VERSION : 0.1
   STRUCT
      dMissionCode : DInt;   // Mission code number
      rgdFireHeadThreshold_cmm : Array[0.."CONST_dNumberOfHeadsCycle"] of DInt;   // Head#x firing threshold [mm/100]
      rgdHeadsPositions_cmm : Array[0.."CONST_dNumberOfHeadsCycle"] of DInt;   // Head#x positions request [mm/100]
      rgxFireHeadON_OFF : Array[0.."CONST_dNumberOfHeadsCycle"] of Bool;   // Head#x firing type request [bit]
      rgxDataToProcessInter : Array[0.."CONST_dNumberOfHeadsCycle"] of Bool;   // Head#x data to process by interrupt
      xGateOpen : Bool;   // Interrupt gate open
      dTargetLineValue_cmm : DInt;   // Virtual target line value [mm/100]
      rgxArmRequest : Array[0.."CONST_dNumberOfHeadsCycle"] of Bool;   // Head#x arming request
      rgdArmRequestTarget_cmm : Array[0.."CONST_dNumberOfHeadsCycle"] of DInt;   // Arm request target virtual [mm/100]
      rgxOilRequest : Array[0.."CONST_dNumberOfHeadsCycle"] of Bool;   // Head#x oil request
      rgdOilRequestTarget_cmm : Array[0.."CONST_dNumberOfHeadsCycle"] of DInt;   // Oil request target virtual [mm/100]
      rgdArmRequestIDMission : Array[0.."CONST_dNumberOfHeadsCycle"] of DInt;   // Arm request ID mission
      rgdOilRequestIDMission : Array[0.."CONST_dNumberOfHeadsCycle"] of DInt;   // Oil request ID mission
   END_STRUCT;
END_TYPE

TYPE "UDT_DataManager_Tank"
VERSION : 0.1
   STRUCT
      dMissionCode : DInt;   // Mission code
      dMissionValue_cmm : DInt;   // Mission value [mm/100]
      rgxFireRequest : Array[0.."CONST_dNumberOfHeadsCycle"] of Bool;   // Head#x fire request
      rgdHeadsPositions_cmm : Array[0.."CONST_dNumberOfHeadsCycle"] of DInt;   // Head#x position request [mm/100]
   END_STRUCT;
END_TYPE

TYPE "UDT_MB_ConnData"
   STRUCT
      IP_OCTET_1 : USInt;
      IP_OCTET_2 : USInt;
      IP_OCTET_3 : USInt;
      IP_OCTET_4 : USInt;
      ConnectID1 : Conn_Ouc;
      ConnectID2 : Conn_Ouc;
      ConnectID3 : Conn_Ouc;
      ConnectID4 : Conn_Ouc;
   END_STRUCT;
END_TYPE

TYPE "UDT_CM_IDEV_FromMainLine"
VERSION : 0.1
   STRUCT
      dSpare1 : Array[0..2] of DInt;
      xCycleON : Bool;   // Cycle ON
      xResetAnomaly : Bool;   // Reset anomaly
      xResetBuffers : Bool;   // Reset buffer
      xGlassBreak : Bool;   // Glass break under the bridge
      xPLCActive0 : Bool;   // PLC Active (0=CPU0, 1=CPU1)
      xPLCActive1 : Bool;   // PLC Active (0=CPU0, 1=CPU1)
      xQLTplate : Bool;   // Quality plate in progress
      xSpare2 : Bool;
      xSpare3 : Bool;
      xSpare4 : Bool;
      xSpare5 : Bool;
      xSpare6 : Bool;
      xSpare7 : Bool;
      xSpare8 : Bool;
      xSpare9 : Bool;
      xSpare10 : Bool;
      xStatusSpare : Array[0..15] of Bool;
      dSpare2 : Array[0..7] of DInt;
      iSpare : Int;
   END_STRUCT;
END_TYPE

TYPE "UDT_CM_IDEV_ToMainLine"
VERSION : 0.1
   STRUCT
      dProcessingIDPlate : DInt;   // Processing ID Plate [Num]
      dSpare1 : DInt;
      dSpare2 : DInt;
      rgxStatus : Array[0..31] of Bool;   // Status heads
      rgdHeadsPositions_cmm : Array[0..15] of DInt;   // Head #x position status
      rgxHeadStatus : Array[0..15] of Bool;   // Head #x enabled
      rgxCuttingStatus : Array[0..15] of Bool;   // Head #x cuuting status
      rgdHeadsPressure : Array[0..15] of DInt;   // Head #x Pressure [mN]
      rgrHeadsSpace : Array[0..15] of Real;   // Head #x Distance [Km]
      iFireOffset_ON : Int;   // All head fire on offset
      iFireOffset_OFF : Int;   // All head fire off offset
      iSpare : Int;
      dSpare : Array[0..7] of DInt;
   END_STRUCT;
   // // rgxStatus[0] : Glass break in progress
   // // rgxStatus[1] : Liftup pushbutton engaged
   // // rgxStatus[2] : Bridge enabled
   // // rgxStatus[3] : Bridge locked
   // // rgxStatus[8] : Fire offset calibration
END_TYPE

TYPE "UDT_CM_RECV_SyncroData"
VERSION : 0.1
   STRUCT
      dMissionID : DInt;   // Mission Identifier
      dSynchroValue_cmm : DInt;   // Counter value in the last synchro [mm/100]
      dSpare : Array[0..7] of DInt;
      xSpare : Array[0..15] of Bool;
      dSpare2 : Array[0..2] of DInt;
      iSpare : Int;
   END_STRUCT;
END_TYPE

TYPE "UDT_CM_RECV_MissionData"
VERSION : 0.1
   STRUCT
      dMissionID : DInt;   // Mission Identifier
      dMissionStart_cmm : DInt;   // Mission counter start [mm/100]
      dMissionEnd_cmm : DInt;   // Mission counter stop [mm/100]
      dTrackingDbNumber : DInt;   // Tracking DB number
      dSpare1 : Array[0..9] of DInt;
      rgxFireRequest : Array[0..31] of Bool;   // Head #x firing request
      rgdHeadsPosition_cmm : Array[0..15] of DInt;   // Head #x position request [mm/100]
      dSpare2 : Array[0..14] of DInt;
   END_STRUCT;
END_TYPE

TYPE "UDT_CM_Manager"
VERSION : 0.1
   STRUCT
      ST_xNewDataReceiveCPU0 : Bool;   // New data receive
      ST_xErrorCPU0 : Bool;   // Error
      ST_xNewSynchCPU0 : Bool;   // New synch
      ST_xNewMissionCPU0 : Bool;   // New mission
      AUX_iDataLenghtCPU0 : Word;   // Data lenght
      AUX_iStateCPU0 : Int;   // Status
      ST_xNewDataReceiveCPU1 : Bool;   // New data receive
      ST_xErrorCPU1 : Bool;   // Error
      ST_xNewSynchCPU1 : Bool;   // New synch
      ST_xNewMissionCPU1 : Bool;   // New mission
      AUX_iDataLenghtCPU1 : Word;   // Data lenght
      AUX_iStateCPU1 : Int;   // Status
      AUX_tmON_ConsumedTimeout : IEC_TIMER;   // Timer ON consumed timeout PLCA
      AUX_rgdHeadMissionIDInProg_Copy : Array[0.."CONST_dNumberOfHeadsCycle"] of DInt;   // Head#x mission ID in progress
      AUX_rgxHeadFiringMissionInProg_Copy : Array[0.."CONST_dNumberOfHeadsCycle"] of Bool;   // Head#x firing mission in progress
      ST_xConsumedTimeout : Bool;   // Consumed message timeout PLCA
      ST_xMissionPacketLost : Bool;   // Mission message packet lost PLC A
      ST_xSyncroPacketLost : Bool;   // Syncro message packet lost PLC A
      ST_MutingFiringOB : Bool;   // Muting Ob30 firing
   END_STRUCT;
END_TYPE

TYPE "UDT_HeadPar"
VERSION : 0.1
   STRUCT
      iAddress : Int;
      iLength : Byte;
      dValue : DInt;
   END_STRUCT;
END_TYPE

TYPE "UDT_AxisParameters"
VERSION : 0.1
   STRUCT
      rgtAxisParameters : Array[0..20] of "UDT_HeadPar";
      dParametersToDownload : DInt;
   END_STRUCT;
END_TYPE

TYPE "UDT_BRCV_FromMainLine"
VERSION : 0.1
   STRUCT
      SyncroData : "UDT_CM_RECV_SyncroData";
      MissionData : "UDT_CM_RECV_MissionData";
   END_STRUCT;
END_TYPE

TYPE "LPD_typeCountFeedbackCh"
VERSION : 0.1
   STRUCT
      countValue : DInt := 16#0000;   // Current count value
      capturedValue : DInt := 16#0000;   // Last Capture value acquired
      measuredValue : Real := 0.0;   // Current measured value
      powerError : Bool := FALSE;   // Incorrect supply voltage L+
      encError : Bool := FALSE;   // Incorrect encoder signal
      ldError : Bool := FALSE;   // Error when loading via control interface
      reserved1 : Bool := FALSE;   // Reserved
      reserved2 : Bool := FALSE;   // Reserved
      reserved3 : Bool := FALSE;   // Reserved
      reserved4 : Bool := FALSE;   // Reserved
      reserved5 : Bool := FALSE;   // Reserved
      commActive : Bool := FALSE;   // Comm active
      resEventAck : Bool := FALSE;   // Reset of event bits active
      ldStsSlot0 : Bool := FALSE;   // Load request for Slot 0 detected and executed (toggling)
      ldStsSlot1 : Bool := FALSE;   // Load request for Slot 1 detected and executed (toggling)
      stsReady : Bool := FALSE;   // Digital on-board I/O started up and parameters assigned
      stsSwGate : Bool := FALSE;   // Software gate status
      reserved7 : Bool := FALSE;   // Reserved
      reserved8 : Bool := FALSE;   // Reserved
      stsDir : Bool := FALSE;   // Direction of last count value change
      stsCount : Bool := FALSE;   // Count pulse detected within last approx. 0.5 s
      stsGate : Bool := FALSE;   // Internal gate status
      stsDQ0 : Bool := FALSE;   // Status HSC DQ0
      stsDQ1 : Bool := FALSE;   // Status HSC DQ1
      stsDI0 : Bool := FALSE;   // Status HSC DI0
      stsDI1 : Bool := FALSE;   // Status HSC DI1
      stsDI2 : Bool := FALSE;   // Status HSC DI2
      eventZero : Bool := FALSE;   // Zero crossing has occurred
      eventUnderflow : Bool := FALSE;   // Underflow has occurred
      eventOverflow : Bool := FALSE;   // Overflow has occurred
      eventCompare0 : Bool := FALSE;   // Comparison event for DQ0 has occurred
      eventCompare1 : Bool := FALSE;   // Comparison event for DQ1 has occurred
      eventSync : Bool := FALSE;   // Synchronization has occurred
      eventCapture : Bool := FALSE;   // Capture event has occurred
      stsMeasInterval : Bool := FALSE;   // Count pulse detected in previous measuring interval
   END_STRUCT;
END_TYPE

TYPE "LPD_typeCountControlCh"
VERSION : 0.1
   STRUCT
      loadValue0 : DWord := 16#0000;   // Load value 0
      loadValue1 : DWord := 16#0000;   // Load value 1
      controlByte : Byte := B#16#00;   // Control byte load value
      swGate : Bool := FALSE;   // Software gate
      tmCtrlDQ0 : Bool := FALSE;   // Enable technological function DQ0
      tmCtrlDQ1 : Bool := FALSE;   // Enable technological function DQ1
      setDQ0 : Bool := FALSE;   // Set DQ0
      setDQ1 : Bool := FALSE;   // Set DQ1
      enSyncUp : Bool := FALSE;   // Enable upward synchronization
      enSyncDown : Bool := FALSE;   // Enable downward synchronization
      enCapture : Bool := FALSE;   // Enable capture function
      resError : Bool := FALSE;   // Reset of saved error states
      resEvent : Bool := FALSE;   // Reset of saved events
      reserved0 : Bool := FALSE;   // Reserved
      reserved1 : Bool := FALSE;   // Reserved
      reserved2 : Bool := FALSE;   // Reserved
      reserved3 : Bool := FALSE;   // Reserved
      reserved4 : Bool := FALSE;   // Reserved
      SetDir : Bool := FALSE;   // Count direction (with encoder without direction signal)
      reserved5 : Byte;   // Reserved
   END_STRUCT;
END_TYPE

// folder: ProfinetDiagnostic

TYPE "TINFO_"
VERSION : 0.1
   STRUCT
      OB_start_info : Array[0..19] of Byte;
      W_20_STATION : Word;
      B22_slave_type : Byte;
      B23_interrupt_type : Byte;
      B24_origination : Byte;
      B25_diag_flag : Byte;
      W26_PN_ID : Word;
      W28_MFG_ID : Word;
      W30_INST_ID : Word;
      other_data : Array[1..70] of Byte;
   END_STRUCT;
END_TYPE

TYPE "AINFO_"
VERSION : 0.1
   STRUCT
      W0_block_type : Word;
      W2_block_length : Word;
      W4_version : Word;
      W6_interrupt_type : Word;
      D8_API : DWord;
      W12_comp_slot_num : Word;
      W14_submodule_slot_num : Word;
      D16_module_ID : DWord;
      D20_submodule_ID : DWord;
      W24_interrupt_specifer : Word;
      Add_W0_format_ID : Word;
      Add_W2_channel_num : Word;
      Add_B4_error_info : Byte;
      Add_B5_data_format : Byte;
      Add_W6_error_type : Word;
      extended_info : Array[34..1431] of Byte;
   END_STRUCT;
END_TYPE

TYPE "PN_Alarm"
VERSION : 0.1
   STRUCT
      word_allarme : Word;
      canale : Int;
   END_STRUCT;
END_TYPE

// folder: (top level)

DATA_BLOCK "PLANT_CONSTANTS"   // DB6
{ S7_Optimized_Access := 'TRUE' }
VERSION : 0.1
   VAR
      CONST_rgxHomeSide : Array[0.."CONST_dNumberOfHeadsCycle"] of Bool;   // Head#x home side [0=Operator Side 1=Opposite operator side]
      CONST_dHOpSideEnc_cmm : Array[0.."CONST_dNumberOfHeadsCycle"] of DInt;   // Operator side head encumbrance [mm/100]
      CONST_dHOppoSideEnc_cmm : Array[0.."CONST_dNumberOfHeadsCycle"] of DInt;   // Opposite operatore side encumbrance [mm/100]
      CONST_rgtHeadPar : Array[0.."CONST_dNumberOfHeadsCycle"] of "UDT_AxisParameters";   // Array of head parameters
   END_VAR
BEGIN
   CONST_rgxHomeSide[0] := false;
   CONST_rgxHomeSide[1] := false;
   CONST_rgxHomeSide[2] := true;
   CONST_rgxHomeSide[3] := true;
END_DATA_BLOCK

DATA_BLOCK "M256_Manag_IDB"   // DB7
{ S7_Optimized_Access := 'TRUE' }
VERSION : 0.1
// stored: InstanceOfName M256_Manager
"M256_Manager"
BEGIN
   M256A_IDB[0].tHMW.dDescentReactTime_ms := 2000;
   M256A_IDB[0].tHMW.dRaiseReactTime_ms := -100;
END_DATA_BLOCK

DATA_BLOCK "Z256_Manager"   // DB9
{ S7_Optimized_Access := 'TRUE' }
VERSION : 0.1
BEGIN
END_DATA_BLOCK

DATA_BLOCK "Z256"   // DB13
{ S7_Optimized_Access := 'TRUE' }
VERSION : 0.1
   VAR
      tmOFF_ResetAlarm : IEC_TIMER;   // Reset alarm
      tmON_24Vdc : IEC_TIMER;   // Presence 24Vdc timer
      tmON_EmergencyOK : IEC_TIMER;   // Emergency OK timer
      ST_xZoneError : Bool;   // Zone error
      ST_xSelectionAutoMode : Bool;   // Automatic mode selection
      ST_xSelectionManualMode : Bool;   // Manual mode selection
      ST_xConditionOKManualMode : Bool;   // Condition OK for manual mode
      ST_xManualModeAccepted : Bool;   // Manual mode accepted
      ST_xAutoModeAccepted : Bool;   // Automatic mode accepted
      ST_xManualModeRequest : Bool;   // Manual mode request
      ST_xFaultsEnabled : Bool;   // Faults enabled
      ST_xZoneEmergency : Bool;   // Cumulative of emergency faults active
      ST_xZoneFaults : Bool;   // Cumulative of zone faults
      ST_xZoneStoppingFaults : Bool;   // Cumulative of zone stopping faults
      ST_xZoneWarnings : Bool;   // Cumulative of zone warning
      ST_xGlassBreak : Bool;   // Glass break under the zone
      ST_xConditionOkBridgeOutProd : Bool;   // Condition OK for bridge out of production
      ST_rgxConditionOkHeadOutProd : Array[0.."CONST_dNumberOfHeadsCycle"] of Bool;   // Condition OK for head out of production
      ST_xCycleON : Bool;   // Zone in cycle ON
      ST_xPLCB_Active : Bool;   // PLC B is active
      OSN_xGateOpen : Bool;   // OSN gate open
      OSR_xGateOpen : Bool;   // OSR gate open
      OS_xGeneralReset : Bool;   // General reset
      OS_xGateOpen : Bool;   // OS gate open
      ON_xGateOpen : Bool;   // ON gate open
      INPUT_xOperatorOverstroke : Bool;   // Operator side head overstroke
      INPUT_xOppoOperatorOverstroke : Bool;   // Opposite operator side head overstroke
      INPUT_xInputCtrlCabinetON : Bool;   // L+.Power supply input control cabinet ON
      INPUT_xInputPowerSupplyON : Bool;   // L+.Input installation power supply ON
      INPUT_xAnomalyPower120_240 : Bool;   // QF.Anomaly power supplies 120 / 240
      INPUT_xPowerSupply24vLogic1 : Bool;   // QF.Power supply 24v logic #1
      INPUT_xPowerSupply24vLogic2 : Bool;   // QF.Power supply 24v logic #2
      INPUT_xPowerSupply24vLogic3 : Bool;   // QF.Power supply 24v logic #3
      INPUT_xPowerSupply24vLogic4 : Bool;   // QF.Power supply 24v logic #4
      INPUT_xPowerSupply24vLogic5 : Bool;   // QF.Power supply 24v logic #5
      INPUT_xLocalEmergencyON : Bool;   // KE.Main emergency ON
      INPUT_xMainEmergencyON : Bool;   // KE.Main emergency ON
      INPUT_xProtSupply36v_1 : Bool;   // QF.Protection power supply 36v #1
      INPUT_xProtSupply36v_2 : Bool;   // QF.Protection power supply motors longitudinal cutting #1
      INPUT_xProtMotorLC_1 : Bool;   // QF.Protection power supply 36v #2
      INPUT_xProtMotorLC_2 : Bool;   // QF.Protection power supply motors longitudinal cutting #2
      INPUT_xProtConditioners : Bool;   // QF.Protection conditioners
      INPUT_xResetLocalEmergency : Bool;   // SB.Reset local emergency
      INPUT_xLocalEmergency_SB1 : Bool;   // SB1.Local emergency
      INPUT_xLocalEmergency_SB2 : Bool;   // SB2.Local emergency
      INPUT_xLocalEmergency_Cabinet : Bool;   // Cabinet.Local emergency
      INPUT_rgxHeadsInProduction : Array[0.."CONST_dNumberOfHeadsCycle"] of Bool;   // SL.Head#x in production
      OUTPUT_xResetLocalEmergency : Bool;   // KM.Reset local emergency
      OUTPUT_xAreaFailure : Bool;   // HL.Cabinet area failure
      OUTPUT_xLocalEmergencyON : Bool;   // HL.Local emergency ON
      OUTPUT_xMachineOutOfOrder : Bool;   // HL.Machine out of order RED
      OUTPUT_xMachineToMaintenance : Bool;   // HL.Machine to maintenance YELLOW
      OUTPUT_xMachineInOrder : Bool;   // HL.Machine in order GREEN
      OUTPUT_xMachineReady : Bool;   // HL.Machine ready WHITE
      OUTPUT_rgxHeadsInProduction : Array[0.."CONST_dNumberOfHeadsCycle"] of Bool;   // HL.Head #x in production
   END_VAR
BEGIN
END_DATA_BLOCK

DATA_BLOCK "Z256_hmi"   // DB14
{ S7_Optimized_Access := 'FALSE' }
VERSION : 0.1
   VAR
      tHMR : Struct   // {[Unit][Scada unit][Low limit][High limit][Access]}
         dCabinetStatus : DInt := 0;   // Cabinet status (0=OK;1=General power alarm;2=Local power alarm) {x|x|x|x|O}
         dZoneMode : DInt := 4;   // Zone modality (1=Manual;4=Automatic;8=Manual request) {x|x|x|x|O}
         xZoneAlarm : Bool := FALSE;   // Zone alarm {x|x|x|x|O}
         xCalibrationsAllowed : Bool := FALSE;   // Calibration function allowed {x|x|x|x|O}
         dProdModeRequest : DInt := 3;   // Production modality request (1=Out of Production 3= In production) {x|x|x|x|O}
         dProdModeActual : DInt := 3;   // Production modality actual (1=Out of production 3=In production 8=Out of production request 9=In production request) {x|x|x|x|O}
         rgdHeadsActualStatus : Array[0.."CONST_dNumberOfHeadsCycle"] of DInt;   // Head status {x|x|x|x|O}
         tManCmd : Struct
            xSpare : Bool := FALSE;
         END_STRUCT;
      END_STRUCT;
      tHMW : Struct   // {[Unit][Scada unit][Low limit][High limit][Access]}
         xFaultsReset : Bool := FALSE;   // Reset faults {x|x|x|x|O}
         xAutoModeReq : Bool := FALSE;   // Automatic mode request {x|x|x|x|O}
         xManModeReq : Bool := FALSE;   // Manual mode request {x|x|x|x|O}
         xOutOfProdReq : Bool := FALSE;   // Bridge out of production request {x|x|x|x|O}
         xInProdReq : Bool := FALSE;   // Bridge in production request {x|x|x|x|O}
         xGeneralReset : Bool := FALSE;   // General reset {x|x|x|x|M}
         xCutOnBreakEnabled : Bool := FALSE;   // Cut during glass break {x|x|x|x|O}
         xMotorsAndCardsInitialize : Bool := FALSE;   // Motors and cards initialize {x|x|x|x|M}
         dNumberOfLites : DInt := 1;   // Calibration. number of lite on calibration {x|x|1|8|M}
         rgdHeadSelected : Array[0.."CONST_dNumberOfHeadsCycle"] of DInt;   // Calibration. head number selected Cut#x{x|x|1|11|M}
         rgdCutWidthTeo_cmm : Array[0.."CONST_dNumberOfHeadsCycle"] of DInt;   // Calibration. cut width Lite #x theorical [mm/100] {mm/100|mm|200|4000|M}
         rgdCutWidthReal_cmm : Array[0.."CONST_dNumberOfHeadsCycle"] of DInt;   // Calibration. cut width real Lite #x [mm/100] {mm/100|mm|200|4000|M}
         xPositionCalibrationRequest : Bool := FALSE;   // Position calibration request {x|x|x|x|M}
         xForceHeadsHoming : Bool := FALSE;   // Force the homing of the heads {x|x|x|x|M}
         xBridgeOffsetCalibrationRequest : Bool := FALSE;   // Bridge offset calibration request {x|x|x|x|M}
         dMoveBridgeOffset_cmm : DInt := 0;   // Calibration. Move all the heads of this offset {mm/100|mm|-100|100|M}
         dPressureScalerOnSample_perc : DInt := 100;   // Pressure scaler during sample plate [%] {%|%|0|100|O}
         rgxHeadEnabled : Array[0.."CONST_dNumberOfHeadsCycle"] of Bool;   // Head enabled/disabled {x|x|x|x|O}
         tManCmd : Struct
            xBrakeEngage : Bool := FALSE;   // Brake engage all heads {x|x|x|x|O}
            xBrakeRelease : Bool := FALSE;   // Brake release all heads {x|x|x|x|O}
         END_STRUCT;
      END_STRUCT;
   END_VAR
BEGIN
   tHMR.rgdHeadsActualStatus[0] := 3;   // Head #x prod. status (1=Out of production 3=In production 8=Out of production request 9=In production request) {x|x|x|x|O}
   tHMR.rgdHeadsActualStatus[1] := 3;   // Head #x prod. status (1=Out of production 3=In production 8=Out of production request 9=In production request) {x|x|x|x|O}
   tHMR.rgdHeadsActualStatus[2] := 3;   // Head #x prod. status (1=Out of production 3=In production 8=Out of production request 9=In production request) {x|x|x|x|O}
   tHMR.rgdHeadsActualStatus[3] := 3;   // Head #x prod. status (1=Out of production 3=In production 8=Out of production request 9=In production request) {x|x|x|x|O}
   tHMW.rgxHeadEnabled[0] := TRUE;   // Head enabled/disabled {x|x|x|x|O}
   tHMW.rgxHeadEnabled[1] := TRUE;   // Head enabled/disabled {x|x|x|x|O}
   tHMW.rgxHeadEnabled[2] := TRUE;   // Head enabled/disabled {x|x|x|x|O}
   tHMW.rgxHeadEnabled[3] := TRUE;   // Head enabled/disabled {x|x|x|x|O}
   // tHMR.rgdHeadsActualStatus[4] : Head #x prod. status (1=Out of production 3=In production 8=Out of production request 9=In production request) {x|x|x|x|O}
   // tHMW.rgdHeadSelected[0] : Calibration. head number selected Cut#x{x|x|1|11|M}
   // tHMW.rgdHeadSelected[1] : Calibration. head number selected Cut#x{x|x|1|11|M}
   // tHMW.rgdHeadSelected[2] : Calibration. head number selected Cut#x{x|x|1|11|M}
   // tHMW.rgdHeadSelected[3] : Calibration. head number selected Cut#x{x|x|1|11|M}
   // tHMW.rgdHeadSelected[4] : Calibration. head number selected Cut#x{x|x|1|11|M}
   // tHMW.rgdCutWidthTeo_cmm[0] : Calibration. cut width Lite #x theorical [mm/100] {mm/100|mm|200|4000|M}
   // tHMW.rgdCutWidthTeo_cmm[1] : Calibration. cut width Lite #x theorical [mm/100] {mm/100|mm|200|4000|M}
   // tHMW.rgdCutWidthTeo_cmm[2] : Calibration. cut width Lite #x theorical [mm/100] {mm/100|mm|200|4000|M}
   // tHMW.rgdCutWidthTeo_cmm[3] : Calibration. cut width Lite #x theorical [mm/100] {mm/100|mm|200|4000|M}
   // tHMW.rgdCutWidthTeo_cmm[4] : Calibration. cut width Lite #x theorical [mm/100] {mm/100|mm|200|4000|M}
   // tHMW.rgdCutWidthReal_cmm[0] : Calibration. cut width real Lite #x [mm/100] {mm/100|mm|200|4000|M}
   // tHMW.rgdCutWidthReal_cmm[1] : Calibration. cut width real Lite #x [mm/100] {mm/100|mm|200|4000|M}
   // tHMW.rgdCutWidthReal_cmm[2] : Calibration. cut width real Lite #x [mm/100] {mm/100|mm|200|4000|M}
   // tHMW.rgdCutWidthReal_cmm[3] : Calibration. cut width real Lite #x [mm/100] {mm/100|mm|200|4000|M}
   // tHMW.rgdCutWidthReal_cmm[4] : Calibration. cut width real Lite #x [mm/100] {mm/100|mm|200|4000|M}
   // tHMW.rgxHeadEnabled[4] : Head enabled/disabled {x|x|x|x|O}
END_DATA_BLOCK

DATA_BLOCK "Z256_alm"   // DB15
{ S7_Optimized_Access := 'FALSE' }
VERSION : 0.1
   VAR
      tE : Struct
         x0 : Bool;   // KE.Main emergency on
         x1 : Bool;   // KE1.Local emergency on
         x2 : Bool;   // Cabinet.Emergency localization
         x3 : Bool;   // SB1.Emergency localization
         x4 : Bool;   // SB2.Emergency localization
         x5 : Bool;
         x6 : Bool;
         x7 : Bool;
         x8 : Bool;
         x9 : Bool;
         x10 : Bool;
         x11 : Bool;
         x12 : Bool;
         x13 : Bool;
         x14 : Bool;
         x15 : Bool;
         x16 : Bool;
         x17 : Bool;
         x18 : Bool;
         x19 : Bool;
         x20 : Bool;
         x21 : Bool;
         x22 : Bool;
         x23 : Bool;
         x24 : Bool;
         x25 : Bool;
         x26 : Bool;
         x27 : Bool;
         x28 : Bool;
         x29 : Bool;
         x30 : Bool;
         x31 : Bool;
      END_STRUCT;
      tS : Struct
         x0 : Bool;   // xB18-3L+.PowerSupplyInputControlCabinetON
         x1 : Bool;   // xB18-7L+.InputInstallationPowerSupplyON"
         x2 : Bool;   // xB11QF1/1D/QF2.Anomaly power supplies 120V
         x3 : Bool;   // xB115KM1/2.AuxiliaryPowerSupplySetIn / xB18QF2.Power supply 24V logic
         x4 : Bool;   // xB410AP1.SafetyOnPanel1" / xB18QF3.Power supply 24V logic
         x5 : Bool;   // xB410AP1.SafetyOnPanel2" / xB20QF2.Power supply 24V logic
         x6 : Bool;   // xB20QF3.Power supply 24V logic
         x7 : Bool;   // xB21QF1.Power supply 24V logic
         x8 : Bool;   // xB140QF2.ProtectionPowerSupplyMotorsYcut"
         x9 : Bool;   // xB41QF2.Protection power supply motors longitudinal cutting
         x10 : Bool;   // xB42QF1.Protection power supply 36V
         x11 : Bool;   // xB42QF2.Protection power supply motors longitudinal cutting
         x12 : Bool;
         x13 : Bool;
         x14 : Bool;
         x15 : Bool;
         x16 : Bool;   // PLCA.Timeout receiving consumed message
         x17 : Bool;   // PLCB.Timeout receiving consumed message
         x18 : Bool;   // PLCA.Mission packet lost
         x19 : Bool;   // PLCB.Mission packet lost
         x20 : Bool;   // PLCA.Syncro packet lost
         x21 : Bool;   // PLCB.Syncro packet lost
         x22 : Bool;   // Syncro.YCut meter gap outside the limits
         x23 : Bool;   // Syncro.Main line meter gap outside the limits
         x24 : Bool;   // Syncro.Timeout receiving meter signal from main line
         x25 : Bool;   // Syncro.Timeout receiving syncro value from mainline
         x26 : Bool;   // Syncro.Unexpected syncro pulse
         x27 : Bool;   // Syncro.Unexpected syncro message
         x28 : Bool;   // Syncro.Machine not syncronized
         x29 : Bool;
         x30 : Bool;
         x31 : Bool;
      END_STRUCT;
      tF : Struct
         x0 : Bool;
         x1 : Bool;
         x2 : Bool;
         x3 : Bool;
         x4 : Bool;
         x5 : Bool;
         x6 : Bool;
         x7 : Bool;
         x8 : Bool;
         x9 : Bool;
         x10 : Bool;
         x11 : Bool;
         x12 : Bool;
         x13 : Bool;
         x14 : Bool;
         x15 : Bool;
         x16 : Bool;
         x17 : Bool;
         x18 : Bool;
         x19 : Bool;
         x20 : Bool;
         x21 : Bool;
         x22 : Bool;
         x23 : Bool;
         x24 : Bool;
         x25 : Bool;
         x26 : Bool;
         x27 : Bool;
         x28 : Bool;
         x29 : Bool;
         x30 : Bool;
         x31 : Bool;
      END_STRUCT;
      tW : Struct
         x0 : Bool;   // PLCA.Timeout receiving consumed message
         x1 : Bool;   // PLCB.Timeout receiving consumed message
         x2 : Bool;   // PLCA.Mission packet lost
         x3 : Bool;   // PLCB.Mission packet lost
         x4 : Bool;   // PLCA.Syncro packet lost
         x5 : Bool;   // PLCB.Syncro packet lost
         x6 : Bool;   // QF.Protection air conditioners
         x7 : Bool;
         x8 : Bool;
         x9 : Bool;
         x10 : Bool;
         x11 : Bool;
         x12 : Bool;
         x13 : Bool;
         x14 : Bool;
         x15 : Bool;
         x16 : Bool;
         x17 : Bool;
         x18 : Bool;
         x19 : Bool;
         x20 : Bool;
         x21 : Bool;
         x22 : Bool;
         x23 : Bool;
         x24 : Bool;
         x25 : Bool;
         x26 : Bool;
         x27 : Bool;
         x28 : Bool;
         x29 : Bool;
         x30 : Bool;
         x31 : Bool;
      END_STRUCT;
   END_VAR
BEGIN
END_DATA_BLOCK

DATA_BLOCK "Encoder"   // DB17
{ S7_Optimized_Access := 'TRUE' }
VERSION : 0.1
   VAR
      ST_xSystemReset : Bool;   // Reset the system
      ST_xMachineSyncronized : Bool;   // Machine is syncronized
      ST_xMeterPulseArrived : Bool;   // Meter pulse arrived
      OS_xError_YCutMeterGapOutsideLimits : Bool;   // Error. YCut meter gap outside the limits
      OS_xError_MainLineMeterGapOutisdeLimits : Bool;   // Error. Main line meter gap outside the limits
      OS_xError_TimeoutReceivingMeterSignal : Bool;   // Error.Timeout receiving meter signal from main line
      OS_xError_TimeoutReceivingSyncroValue : Bool;   // Error.Timeout receiving syncro value from mainline
      OS_xError_UnexpectedSyncroPulse : Bool;   // Error.Unexpected syncro pulse
      OS_xError_UnexpectedSyncroMessage : Bool;   // Error.Unexpected syncro message
      OSR_xMeterPulse : Bool;   // OSR Meter pulse
      OS_xMeterPulse : Bool;   // OS Meter pulse
      PH_WaitFirstMeter : Bool;   // Waiting first meter pulse
      PH_EndWaitFirstMeter : Bool;   // End waiting first meter pulse
      PH_WaitFirstMeterDataFromMain : Bool;   // Waiting first meter data from main
      PH_EndWaitFirstMeterDataFromMain : Bool;   // End waiting first meter data from main
      PH_WaitMeterPulse : Bool;   // Waiting meter pulse
      PH_EndWaitMeterPulse : Bool;   // End waiting meter pulse
      PH_WaitMeterDataFromMain : Bool;   // Wait meter data from main line
      PH_EndWaitMeterDataFromMain : Bool;   // End wait meter data from main line
      AUX_dActualEncoderValue_cmm : DInt;   // Actual encoder pulse value [mm/100]
      AUX_dActualSpeedValue_cmm_min : DInt;   // Actual lehr speed [cmm/min]
      AUX_dActualSpeedValue_cmm_s : DInt;   // Actual lehr speed [cmm/s]
      AUX_rActualSpeedValue_cmm_ms : Real;   // Actual lehr speed [mm/100 /ms]
      AUX_xNewSyncroReceived : Bool;   // New syncro received from master
      AUX_dNewSyncroValue_cmm : DInt;   // New value of syncro received [mm/100]
      AUX_dLastMainLineValue_cmm : DInt;   // Last main line value syncro [mm/100]
      AUX_dLastStoredSyncroValue_cmm : DInt;   // Last stored syncro value [mm/100]
      AUX_dSyncroGapMainLine_cmm : DInt;   // Syncro gap beetween main line and ycut [mm/100]
      AUX_dMissingSyncroCounter : DInt;   // Missing syncro counter
      AUX_dMeterPulseValue_count : DInt;   // Meter pulse value
      INPUT_dEncoderCounter_count : DInt;   // Encoder counter [count]
      INPUT_dFrequencyCounter_Hz : DInt;   // Frequency counter [Hz]
      INPUT_xMeterPulseArrived : Bool;   // Meter pulse arrived
      INPUT_dMeterPulseValue_count : DInt;   // Meter pulse value [count]
      INPUT_xResetEventAcknowledge : Bool;   // Reset event bit active
      OUTPUT_xCounterEnable : Bool;   // Enable card counter
      OUTPUT_xCounterReset : Bool;   // Card counter reset
      OUTPUT_xResetMeterPulse : Bool;   // Reset meter pulse
      AUX_tmOFFResetMeter : IEC_TIMER;   // Retain meter pulse
      AUX_tmOFFRetainCardReset : IEC_TIMER;   // Retain encoder card reset
   END_VAR
BEGIN
END_DATA_BLOCK

DATA_BLOCK "M256_Manag_Init"   // DB20
{ S7_Optimized_Access := 'TRUE' }
VERSION : 0.1
// stored: InstanceOfName M256_Manager
"M256_Manager"
BEGIN
END_DATA_BLOCK

// folder: 07_ArrayScada

DATA_BLOCK "DB_Z256_Scada"   // DB2010
{ S7_Optimized_Access := 'FALSE' }
VERSION : 0.1
   VAR
      tAlm : Struct   // HMI Alarms
         tE : Struct
            x0 : Bool;   // KE.Main emergency on
            x1 : Bool;   // KE1.Local emergency on
            x2 : Bool;   // Cabinet.Emergency localization
            x3 : Bool;   // SB1.Emergency localization
            x4 : Bool;   // SB2.Emergency localization
            x5 : Bool;
            x6 : Bool;
            x7 : Bool;
            x8 : Bool;
            x9 : Bool;
            x10 : Bool;
            x11 : Bool;
            x12 : Bool;
            x13 : Bool;
            x14 : Bool;
            x15 : Bool;
            x16 : Bool;
            x17 : Bool;
            x18 : Bool;
            x19 : Bool;
            x20 : Bool;
            x21 : Bool;
            x22 : Bool;
            x23 : Bool;
            x24 : Bool;
            x25 : Bool;
            x26 : Bool;
            x27 : Bool;
            x28 : Bool;
            x29 : Bool;
            x30 : Bool;
            x31 : Bool;
         END_STRUCT;
         tS : Struct
            tS0 : Struct
               x0 : Bool;   // xB18-3L+.PowerSupplyInputControlCabinetON
               x1 : Bool;   // xB18-7L+.InputInstallationPowerSupplyON"
               x2 : Bool;   // xB11QF1/1D/QF2.Anomaly power supplies 120V
               x3 : Bool;   // xB115KM1/2.AuxiliaryPowerSupplySetIn / xB18QF2.Power supply 24V logic
               x4 : Bool;   // xB410AP1.SafetyOnPanel1" / xB18QF3.Power supply 24V logic
               x5 : Bool;   // xB410AP1.SafetyOnPanel2" / xB20QF2.Power supply 24V logic
               x6 : Bool;   // xB20QF3.Power supply 24V logic
               x7 : Bool;   // xB21QF1.Power supply 24V logic
               x8 : Bool;   // xB140QF2.ProtectionPowerSupplyMotorsYcut" / xB41QF1.ProtectionPowerSupplyMotorsYcut 1-4
               x9 : Bool;   // xB41QF2.Protection power supply motors longitudinal cutting / xB41QF2.Protection power supply 36V motors longitudinal cutting 1-4
               x10 : Bool;   // xB42QF1.Protection power supply 36V / xB42QF1.ProtectionPowerSupplyMotorsYcut 5-8
               x11 : Bool;   // xB42QF2.Protection power supply motors longitudinal cutting / xB42QF2.Protection power supply 36V motors longitudinal cutting 5-8
               x12 : Bool;
               x13 : Bool;
               x14 : Bool;
               x15 : Bool;
               x16 : Bool;   // PLCA.Timeout receiving consumed message
               x17 : Bool;   // PLCB.Timeout receiving consumed message
               x18 : Bool;   // PLCA.Mission packet lost
               x19 : Bool;   // PLCB.Mission packet lost
               x20 : Bool;   // PLCA.Syncro packet lost
               x21 : Bool;   // PLCB.Syncro packet lost
               x22 : Bool;   // Syncro.YCut meter gap outside the limits
               x23 : Bool;   // Syncro.Main line meter gap outside the limits
               x24 : Bool;   // Syncro.Timeout receiving meter signal from main line
               x25 : Bool;   // Syncro.Timeout receiving syncro value from mainline
               x26 : Bool;   // Syncro.Unexpected syncro pulse
               x27 : Bool;   // Syncro.Unexpected syncro message
               x28 : Bool;   // Syncro.Machine not syncronized
               x29 : Bool;
               x30 : Bool;
               x31 : Bool;
            END_STRUCT;
            tS1 : Struct
               x0 : Bool;
               x1 : Bool;   // Syncro.YCut meter gap outside the limits
               x2 : Bool;
               x3 : Bool;
               x4 : Bool;
               x5 : Bool;
               x6 : Bool;
               x7 : Bool;
               x8 : Bool;   // xB21QF1.Power supply 24V logic
               x9 : Bool;
               x10 : Bool;   // Syncro.Main line meter gap outside the limits
               x11 : Bool;
               x12 : Bool;
               x13 : Bool;
               x14 : Bool;
               x15 : Bool;
               x16 : Bool;
               x17 : Bool;
               x18 : Bool;
               x19 : Bool;
               x20 : Bool;
               x21 : Bool;
               x22 : Bool;
               x23 : Bool;
               x24 : Bool;
               x25 : Bool;
               x26 : Bool;
               x27 : Bool;
               x28 : Bool;
               x29 : Bool;
               x30 : Bool;
               x31 : Bool;
            END_STRUCT;
            tS2 : Struct
               x0 : Bool;
               x1 : Bool;   // Syncro.YCut meter gap outside the limits
               x2 : Bool;
               x3 : Bool;
               x4 : Bool;
               x5 : Bool;
               x6 : Bool;
               x7 : Bool;
               x8 : Bool;   // xB21QF1.Power supply 24V logic
               x9 : Bool;
               x10 : Bool;   // Syncro.Main line meter gap outside the limits
               x11 : Bool;
               x12 : Bool;
               x13 : Bool;
               x14 : Bool;
               x15 : Bool;
               x16 : Bool;
               x17 : Bool;
               x18 : Bool;
               x19 : Bool;
               x20 : Bool;
               x21 : Bool;
               x22 : Bool;
               x23 : Bool;
               x24 : Bool;
               x25 : Bool;
               x26 : Bool;
               x27 : Bool;
               x28 : Bool;
               x29 : Bool;
               x30 : Bool;
               x31 : Bool;
            END_STRUCT;
            tS3 : Struct
               x0 : Bool;
               x1 : Bool;   // Syncro.YCut meter gap outside the limits
               x2 : Bool;
               x3 : Bool;
               x4 : Bool;
               x5 : Bool;
               x6 : Bool;
               x7 : Bool;
               x8 : Bool;   // xB21QF1.Power supply 24V logic
               x9 : Bool;
               x10 : Bool;   // Syncro.Main line meter gap outside the limits
               x11 : Bool;
               x12 : Bool;
               x13 : Bool;
               x14 : Bool;
               x15 : Bool;
               x16 : Bool;
               x17 : Bool;
               x18 : Bool;
               x19 : Bool;
               x20 : Bool;
               x21 : Bool;
               x22 : Bool;
               x23 : Bool;
               x24 : Bool;
               x25 : Bool;
               x26 : Bool;
               x27 : Bool;
               x28 : Bool;
               x29 : Bool;
               x30 : Bool;
               x31 : Bool;
            END_STRUCT;
         END_STRUCT;
         tF : Struct
            x0 : Bool;
            x1 : Bool;
            x2 : Bool;
            x3 : Bool;
            x4 : Bool;
            x5 : Bool;
            x6 : Bool;
            x7 : Bool;
            x8 : Bool;
            x9 : Bool;
            x10 : Bool;
            x11 : Bool;
            x12 : Bool;
            x13 : Bool;
            x14 : Bool;
            x15 : Bool;
            x16 : Bool;
            x17 : Bool;
            x18 : Bool;
            x19 : Bool;
            x20 : Bool;
            x21 : Bool;
            x22 : Bool;
            x23 : Bool;
            x24 : Bool;
            x25 : Bool;
            x26 : Bool;
            x27 : Bool;
            x28 : Bool;
            x29 : Bool;
            x30 : Bool;
            x31 : Bool;
         END_STRUCT;
         tW : Struct
            x0 : Bool;   // PLCA.Timeout receiving consumed message
            x1 : Bool;   // PLCB.Timeout receiving consumed message
            x2 : Bool;   // PLCA.Mission packet lost
            x3 : Bool;   // PLCB.Mission packet lost
            x4 : Bool;   // PLCA.Syncro packet lost
            x5 : Bool;   // PLCB.Syncro packet lost
            x6 : Bool;   // QF.Protection air conditioners
            x7 : Bool;
            x8 : Bool;
            x9 : Bool;
            x10 : Bool;
            x11 : Bool;
            x12 : Bool;
            x13 : Bool;
            x14 : Bool;
            x15 : Bool;
            x16 : Bool;
            x17 : Bool;
            x18 : Bool;
            x19 : Bool;
            x20 : Bool;
            x21 : Bool;
            x22 : Bool;
            x23 : Bool;
            x24 : Bool;
            x25 : Bool;
            x26 : Bool;
            x27 : Bool;
            x28 : Bool;
            x29 : Bool;
            x30 : Bool;
            x31 : Bool;
         END_STRUCT;
      END_STRUCT;
      tHMR : Struct   // HMI Read
         xCalibrationsAllowed : Bool := FALSE;   // Calibration function allowed {x|x|x|x|O}
         xSpare1 : Bool;
         xSpare2 : Bool;
         xSpare3 : Bool;
         xSpare4 : Bool;
         xSpare5 : Bool;
         xSpare6 : Bool;
         xSpare7 : Bool;
         xSpare8 : Bool;
         xSpare9 : Bool;
         xSpare10 : Bool;
         xSpare11 : Bool;
         xSpare12 : Bool;
         xSpare13 : Bool;
         xSpare14 : Bool;
         xZoneAlarm : Bool := FALSE;   // Zone alarm {X|X|X|X|O}
         xSpare16 : Bool;
         xSpare17 : Bool;
         xSpare18 : Bool;
         xSpare19 : Bool;
         xSpare20 : Bool;
         xSpare21 : Bool;
         xSpare22 : Bool;
         xSpare23 : Bool;
         xSpare24 : Bool;
         xSpare25 : Bool;
         xSpare26 : Bool;
         xSpare27 : Bool;
         xSpare28 : Bool;
         xSpare29 : Bool;
         xSpare30 : Bool;
         xSpare31 : Bool;
         xSpare : Array[0..15] of Bool;
         iSpare0 : Int;
         iSpare1 : Int;
         iSpare2 : Int;
         iSpare3 : Int;
         iSpare4 : Int;
         iSpare5 : Int;
         iSpare6 : Int;
         iSpare7 : Int;
         iSpare8 : Int;
         iSpare9 : Int;
         iSpare10 : Int;
         iSpare11 : Int;
         iSpare12 : Int;
         iSpare13 : Int;
         iSpare14 : Int;
         iSpare15 : Int;
         iSpare16 : Int;
         dZoneMode : DInt := 4;   // Zone modality (1=Manual;4=Automatic;8=Manual request) {x|x|x|x|O}
         dZoneState : DInt := 1024;   // Zone status (1=CycleON 2=StopCyc 4=CycleReq 8=StopReq 1024=E-Stop) {X|X|X|X|O} / HMI Alarms
         dCabinetStatusMCC : DInt := 1;   // Cabinet status MCC1256B (1=OK;2=General power alarm;3=Local power alarm) {X|X|X|X|O} / HMI Write
         dProdModeRequest : DInt := 3;   // Production modality request (1=Out of Production 3= In production) {x|x|x|x|O}
         dProdModeActual : DInt := 3;   // Production modality actual (1=Out of production 3=In production 8=Out of production request 9=In production request) {x|x|x|x|O}
         dSpare5 : DInt;
         "rgdHeadsActualStatus[0]" : DInt := 3;   // Head #1 prod. status (1=Out of production 3=In production 8=Out of production request 9=In production request) {x|x|x|x|O}
         "rgdHeadsActualStatus[1]" : DInt := 3;   // Head #2 prod. status (1=Out of production 3=In production 8=Out of production request 9=In production request) {x|x|x|x|O}
         "rgdHeadsActualStatus[2]" : DInt := 3;   // Head #3 prod. status (1=Out of production 3=In production 8=Out of production request 9=In production request) {x|x|x|x|O}
         "rgdHeadsActualStatus[3]" : DInt := 3;   // Head #4 prod. status (1=Out of production 3=In production 8=Out of production request 9=In production request) {x|x|x|x|O}
         "rgdHeadsActualStatus[4]" : DInt;   // Head #5 prod. status (1=Out of production 3=In production 8=Out of production request 9=In production request) {x|x|x|x|O}
         "rgdHeadsActualStatus[5]" : DInt;   // Head #6 prod. status (1=Out of production 3=In production 8=Out of production request 9=In production request) {x|x|x|x|O}
         "rgdHeadsActualStatus[6]" : DInt;   // Head #7 prod. status (1=Out of production 3=In production 8=Out of production request 9=In production request) {x|x|x|x|O}
         "rgdHeadsActualStatus[7]" : DInt;   // Head #8 prod. status (1=Out of production 3=In production 8=Out of production request 9=In production request) {x|x|x|x|O}
         dSpare14 : DInt;
         dSpare15 : DInt;
         dSpare : Array[0..15] of DInt;
         rSpare0 : Real;
         rSpare1 : Real;
         rSpare2 : Real;
         rSpare3 : Real;
         rSpare4 : Real;
         rSpare5 : Real;
         rSpare6 : Real;
         rSpare7 : Real;
         rSpare8 : Real;
         tManCmd : Struct
            xSpare0 : Bool;
            xSpare1 : Bool;
            xSpare2 : Bool;
            xSpare3 : Bool;
            xSpare4 : Bool;
            xSpare5 : Bool;
            xSpare6 : Bool;
            xSpare7 : Bool;
            xSpare8 : Bool;
            xSpare9 : Bool;
            xSpare10 : Bool;
            xSpare11 : Bool;
            xSpare12 : Bool;
            xSpare13 : Bool;
            xSpare14 : Bool;
            xSpare15 : Bool;
            xSpare : Array[0..15] of Bool;
         END_STRUCT;
      END_STRUCT;
      tHMW : Struct   // HMI Write
         xAutoModeReq : Bool := FALSE;   // Automatic mode request {x|x|x|x|O}
         xManModeReq : Bool := FALSE;   // Manual mode request {x|x|x|x|O}
         xOutOfProdReq : Bool := FALSE;   // Bridge out of production request {x|x|x|x|O}
         xInProdReq : Bool := FALSE;   // Bridge in production request {x|x|x|x|O}
         xCutOnBreakEnabled : Bool := FALSE;   // Cut during glass break {x|x|x|x|O}
         xMotorsAndCardsInitialize : Bool := FALSE;   // Motors and cards initialize {x|x|x|x|M}
         xForceHeadsHoming : Bool := FALSE;   // Force the homing of the heads {x|x|x|x|M}
         xPositionCalibrationRequest : Bool := FALSE;   // Position calibration request {x|x|x|x|M}
         xBridgeOffsetCalibrationRequest : Bool := FALSE;   // Bridge offset calibration request {x|x|x|x|M}
         xSpare9 : Bool;
         xSpare10 : Bool;
         xSpare11 : Bool;
         xSpare12 : Bool;
         xSpare13 : Bool;
         xGeneralReset : Bool := FALSE;   // General reset {X|X|X|X|M}
         xFaultsReset : Bool := FALSE;   // Reset faults {X|X|X|X|O}
         xHeadEnabled_1 : Bool := TRUE;   // Head #1 enabled/disabled {x|x|x|x|O}
         xHeadEnabled_2 : Bool := TRUE;   // Head #2 enabled/disabled {x|x|x|x|O}
         xHeadEnabled_3 : Bool := TRUE;   // Head #3 enabled/disabled {x|x|x|x|O}
         xHeadEnabled_4 : Bool := TRUE;   // Head #4 enabled/disabled {x|x|x|x|O}
         xHeadEnabled_5 : Bool := TRUE;   // Head #5 enabled/disabled {x|x|x|x|O}
         xHeadEnabled_6 : Bool := TRUE;   // Head #6 enabled/disabled {x|x|x|x|O}
         xHeadEnabled_7 : Bool := TRUE;   // Head #7 enabled/disabled {x|x|x|x|O}
         xHeadEnabled_8 : Bool := TRUE;   // Head #8 enabled/disabled {x|x|x|x|O}
         xSpare24 : Bool;
         xSpare25 : Bool;
         xSpare26 : Bool;
         xSpare27 : Bool;
         xSpare28 : Bool;
         xSpare29 : Bool;
         xSpare30 : Bool;
         xSpare31 : Bool;
         xSpare : Array[0..15] of Bool;
         iSpare0 : Int;
         iSpare1 : Int;
         iSpare2 : Int;
         iSpare3 : Int;
         iSpare4 : Int;
         iSpare5 : Int;
         iSpare6 : Int;
         iSpare7 : Int;
         iSpare8 : Int;
         iSpare9 : Int;
         iSpare10 : Int;
         iSpare11 : Int;
         iSpare12 : Int;
         iSpare13 : Int;
         iSpare14 : Int;
         iSpare15 : Int;
         iSpare16 : Int;
         dNumberOfLites : DInt := 1;   // Calibration. number of lite on calibration {x|x|1|8|M}
         dMoveBridgeOffset_cmm : DInt := 0;   // Calibration. Move all the heads of this offset {mm/100|mm|-100|100|M}
         dPressureScalerOnSample_perc : DInt := 100;   // Pressure scaler during sample plate [%] {%|%|0|100|O}
         dSpare3 : DInt;
         dSpare4 : DInt;
         dSpare5 : DInt;
         dSpare6 : DInt;
         dSpare7 : DInt;
         dHead_Selected_1 : DInt;   // Calibration. head number selected Cut1 {x|x|1|11|M}
         dHead_Selected_2 : DInt;   // Calibration. head number selected Cut2 {x|x|1|11|M}
         dHead_Selected_3 : DInt;   // Calibration. head number selected Cut3{x|x|1|11|M}
         dHead_Selected_4 : DInt;   // Calibration. head number selected Cut4{x|x|1|11|M}
         dHead_Selected_5 : DInt;   // Calibration. head number selected Cut5{x|x|1|11|M}
         dHead_Selected_6 : DInt;   // Calibration. head number selected Cut6{x|x|1|11|M}
         dHead_Selected_7 : DInt;   // Calibration. head number selected Cut7{x|x|1|11|M}
         dHead_Selected_8 : DInt;   // Calibration. head number selected Cut8{x|x|1|11|M}
         dCutWidthTeo_cmm_1 : DInt;   // Calibration. cut width Lite 1 theorical [mm/100] {mm/100|mm|200|4000|M}
         dCutWidthTeo_cmm_2 : DInt;   // Calibration. cut width Lite 2 theorical [mm/100] {mm/100|mm|200|4000|M}
         dCutWidthTeo_cmm_3 : DInt;   // Calibration. cut width Lite 3 theorical [mm/100] {mm/100|mm|200|4000|M}
         dCutWidthTeo_cmm_4 : DInt;   // Calibration. cut width Lite 4 theorical [mm/100] {mm/100|mm|200|4000|M}
         dCutWidthTeo_cmm_5 : DInt;   // Calibration. cut width Lite 5 theorical [mm/100] {mm/100|mm|200|4000|M}
         dCutWidthTeo_cmm_6 : DInt;   // Calibration. cut width Lite 6 theorical [mm/100] {mm/100|mm|200|4000|M}
         dCutWidthTeo_cmm_7 : DInt;   // Calibration. cut width Lite 7 theorical [mm/100] {mm/100|mm|200|4000|M}
         dCutWidthTeo_cmm_8 : DInt;   // Calibration. cut width Lite 8 theorical [mm/100] {mm/100|mm|200|4000|M}
         dCutWidthReal_cmm_1 : DInt;   // Calibration. cut width Lite 1 real [mm/100] {mm/100|mm|200|4000|M}
         dCutWidthReal_cmm_2 : DInt;   // Calibration. cut width Lite 2 real [mm/100] {mm/100|mm|200|4000|M}
         dCutWidthReal_cmm_3 : DInt;   // Calibration. cut width Lite 3 real [mm/100] {mm/100|mm|200|4000|M}
         dCutWidthReal_cmm_4 : DInt;   // Calibration. cut width Lite 4 real [mm/100] {mm/100|mm|200|4000|M}
         dCutWidthReal_cmm_5 : DInt;   // Calibration. cut width Lite 5 real [mm/100] {mm/100|mm|200|4000|M}
         dCutWidthReal_cmm_6 : DInt;   // Calibration. cut width Lite 6 real [mm/100] {mm/100|mm|200|4000|M}
         dCutWidthReal_cmm_7 : DInt;   // Calibration. cut width Lite 7 real [mm/100] {mm/100|mm|200|4000|M}
         dCutWidthReal_cmm_8 : DInt;   // Calibration. cut width Lite 8 real [mm/100] {mm/100|mm|200|4000|M}
         dSpare32 : DInt;
         dSpare33 : DInt;
         dSpare34 : DInt;
         dSpare35 : DInt;
         dSpare36 : DInt;
         dSpare37 : DInt;
         dSpare38 : DInt;
         dSpare39 : DInt;
         dSpare : Array[0..19] of DInt;
         rSpare0 : Real;
         rSpare1 : Real;
         rSpare2 : Real;
         rSpare3 : Real;
         rSpare4 : Real;
         rSpare5 : Real;
         rSpare6 : Real;
         rSpare7 : Real;
         rSpare8 : Real;
         tManCmd : Struct
            xBrakeEngage : Bool := FALSE;   // Brake engage all heads {x|x|x|x|O}
            xBrakeRelease : Bool := FALSE;   // Brake release all heads {x|x|x|x|O}
            xSpare2 : Bool;
            xSpare3 : Bool;
            xSpare4 : Bool;
            xSpare5 : Bool;
            xSpare6 : Bool;
            xSpare7 : Bool;
            xSpare8 : Bool;
            xSpare9 : Bool;
            xSpare10 : Bool;
            xSpare11 : Bool;
            xSpare12 : Bool;
            xSpare13 : Bool;
            xSpare14 : Bool;
            xSpare15 : Bool;
            xSpare16 : Bool;
            xSpare17 : Bool;
            xSpare18 : Bool;
            xSpare19 : Bool;
            xSpare20 : Bool;
            xSpare21 : Bool;
            xSpare22 : Bool;
            xSpare23 : Bool;
            xSpare24 : Bool;
            xSpare25 : Bool;
            xSpare26 : Bool;
            xSpare27 : Bool;
            xSpare28 : Bool;
            xSpare29 : Bool;
            xSpare30 : Bool;
            xSpare31 : Bool;
         END_STRUCT;
      END_STRUCT;
   END_VAR
BEGIN
END_DATA_BLOCK

